(* Logix 5000 project; controller PLC_MCC1300_75F1 vendor 1 type 14 code 166 rev 32.11; software revision 32.04; part 79 of 83 *)
(* tags used below, declared in another part *)
   AUX_xInitialize : BOOL;
   GP_NetDiag : GP_NetworkDiag;
   GP_OB_InitializeDiag : GP_OB_Initialize;
   GP_OB_InitializeDiag_STC : GP_OB_Initialize_STC;
   GP_OB_InitializeMain : GP_OB_Initialize;
   M302SpeedUp : MAC_SpeedUp;
   M307A_M1_DR : AXIS_CIP_DRIVE;
   M307A_M2_DR : AXIS_CIP_DRIVE;
   M307A_M3_DR : AXIS_CIP_DRIVE;
   M351_ALM : MAC_Conveyor_ALM;
   M352_ALM : MAC_Conveyor_ALM;
   M353_ALM : MAC_Conveyor_ALM;
   MCC1300_rgtDiagModule_HMI : GP_NetworkDiag_v1[90];
   TMP_dDirection : DINT;
   TMP_dTarget : DINT;
   TMP_rAcc : REAL;
   TMP_rDec : REAL;
   TMP_rSpeed : REAL;
   Z300_Conveyor : UDT_StandConv[29];
   Z300_Conveyor_IN_MOTION : MAC_Conveyor_ZC_IN_MOTION[29];
   Z300_Conveyor_OUT_MOTION : MAC_Conveyor_ZC_OUT_MOTION[29];
   Z301 : MAC_Zone_ML;
   Z900 : MAC_Zone;
   Z900_HMR : MAC_Zone_HMR;
   Z900_HMW : MAC_Zone_HMW;
(* MainProgram, continued *)

   // #####_HMI_STATUSES_#####
   40: NOP();
   41: XIC(Z900.ST_xZoneError)OTE(Z900_HMR.xZoneAlarm);
   42: XIC(Z900.ST_xCleaningAccepted)OTE(Z900_HMR.xCleaningEnabled);
   43: [MOV(0,Z900_HMR.dCabinetState1) ,[XIC(M351_ALM.rgxStoppingFault_M[0].1) ,XIC(M352_ALM.rgxStoppingFault_M[0].1) ,XIC(M353_ALM.rgxStoppingFault_M[0].1) ] MOV(2,Z900_HMR.dCabinetState1) ,XIC(Z301.OUTPUT_xMCCSafetyLamp) MOV(1,Z900_HMR.dCabinetState1) ];
   44: [XIC(Z900.ST_xManualModeAccepted) MOV(1,Z900_HMR.dZoneMode) ,XIC(Z900.ST_xAutoModeAccepted) MOV(4,Z900_HMR.dZoneMode) ,XIC(Z900.ST_xManualModeRequest) MOV(8,Z900_HMR.dZoneMode) ];
   45: [MOV(2,Z900_HMR.dZoneState) ,XIC(Z900.ST_xStartCycleRequest) XIO(Z900.ST_xCycleON) MOV(4,Z900_HMR.dZoneState) ,XIC(Z900.ST_xCycleON) MOV(1,Z900_HMR.dZoneState) ,XIC(Z900.ST_xStopCycleRequest) MOV(8,Z900_HMR.dZoneState) ,XIO(Z301.INPUT_xMainEmergencyON) MOV(1024,Z900_HMR.dZoneState) ];
   46: [XIC(Z900.ST_xCleaningAccepted) MOV(1,Z900_HMR.dCleaningState) ,XIO(Z900.ST_xCleaningAccepted) MOV(2,Z900_HMR.dCleaningState) ,XIC(Z900.ST_xReqCleaning) XIO(Z900.ST_xCleaningAccepted) MOV(4,Z900_HMR.dCleaningState) ];
   47: [XIC(Z900_HMW.rgxMan.0) OTE(Z900_HMR.rgxMan.0) ,XIC(Z900_HMW.rgxMan.1) OTE(Z900_HMR.rgxMan.1) ];
END_ROUTINE
END_PROGRAM

PROGRAM Modules   (* main routine Main *)

ROUTINE Main   (* ladder *)
   0: GP_OB_Initialize(GP_OB_InitializeDiag,GP_OB_InitializeDiag_STC,AUX_xInitialize);
   1: GP_NetworkDiag(GP_NetDiag,GP_OB_InitializeDiag,ETH_MCC1300,MCC1300_rgtDiagModule_HMI[0]);
   2: GP_NetworkDiag(GP_NetDiag,GP_OB_InitializeDiag,ETH_M2,MCC1300_rgtDiagModule_HMI[1]);
   3: GP_NetworkDiag(GP_NetDiag,GP_OB_InitializeDiag,TD5680AP1,MCC1300_rgtDiagModule_HMI[5]);
   4: GP_NetworkDiag(GP_NetDiag,GP_OB_InitializeDiag,M3683AP1,MCC1300_rgtDiagModule_HMI[6]);
   5: GP_NetworkDiag(GP_NetDiag,GP_OB_InitializeDiag,E152AP1,MCC1300_rgtDiagModule_HMI[7]);
   6: GP_NetworkDiag(GP_NetDiag,GP_OB_InitializeDiag,RIOM13,MCC1300_rgtDiagModule_HMI[8]);
   7: GP_NetworkDiag(GP_NetDiag,GP_OB_InitializeDiag,M3AZ01,MCC1300_rgtDiagModule_HMI[11]);
   8: GP_NetworkDiag(GP_NetDiag,GP_OB_InitializeDiag,M3AZ02,MCC1300_rgtDiagModule_HMI[12]);
   9: GP_NetworkDiag(GP_NetDiag,GP_OB_InitializeDiag,M3AZ03,MCC1300_rgtDiagModule_HMI[13]);
   10: GP_NetworkDiag(GP_NetDiag,GP_OB_InitializeDiag,M3AZ04,MCC1300_rgtDiagModule_HMI[14]);
   11: GP_NetworkDiag(GP_NetDiag,GP_OB_InitializeDiag,M3AZ05,MCC1300_rgtDiagModule_HMI[15]);
   12: GP_NetworkDiag(GP_NetDiag,GP_OB_InitializeDiag,M3AZ06,MCC1300_rgtDiagModule_HMI[16]);
   13: GP_NetworkDiag(GP_NetDiag,GP_OB_InitializeDiag,M3AZ07,MCC1300_rgtDiagModule_HMI[17]);
   14: GP_NetworkDiag(GP_NetDiag,GP_OB_InitializeDiag,M3AZ08,MCC1300_rgtDiagModule_HMI[18]);
   15: GP_NetworkDiag(GP_NetDiag,GP_OB_InitializeDiag,M3AZ09,MCC1300_rgtDiagModule_HMI[19]);
   16: GP_NetworkDiag(GP_NetDiag,GP_OB_InitializeDiag,M3AZ10,MCC1300_rgtDiagModule_HMI[20]);
   17: GP_NetworkDiag(GP_NetDiag,GP_OB_InitializeDiag,TDKAZ00N,MCC1300_rgtDiagModule_HMI[21]);
   18: GP_NetworkDiag(GP_NetDiag,GP_OB_InitializeDiag,TDKAZ00S,MCC1300_rgtDiagModule_HMI[22]);
   19: GP_NetworkDiag(GP_NetDiag,GP_OB_InitializeDiag,TDKAZ01N,MCC1300_rgtDiagModule_HMI[23]);
   20: GP_NetworkDiag(GP_NetDiag,GP_OB_InitializeDiag,TDKAZ01S,MCC1300_rgtDiagModule_HMI[24]);
   21: GP_NetworkDiag(GP_NetDiag,GP_OB_InitializeDiag,TDKAZ02N,MCC1300_rgtDiagModule_HMI[25]);
   22: GP_NetworkDiag(GP_NetDiag,GP_OB_InitializeDiag,TDKAZ02S,MCC1300_rgtDiagModule_HMI[26]);
   23: GP_NetworkDiag(GP_NetDiag,GP_OB_InitializeDiag,TDKAZ03N,MCC1300_rgtDiagModule_HMI[27]);
   24: GP_NetworkDiag(GP_NetDiag,GP_OB_InitializeDiag,TDKAZ03S,MCC1300_rgtDiagModule_HMI[28]);
   25: GP_NetworkDiag(GP_NetDiag,GP_OB_InitializeDiag,TDKAZ04N,MCC1300_rgtDiagModule_HMI[29]);
   26: GP_NetworkDiag(GP_NetDiag,GP_OB_InitializeDiag,TDKAZ04S,MCC1300_rgtDiagModule_HMI[30]);
   27: GP_NetworkDiag(GP_NetDiag,GP_OB_InitializeDiag,TDKAZ05N,MCC1300_rgtDiagModule_HMI[31]);
   28: GP_NetworkDiag(GP_NetDiag,GP_OB_InitializeDiag,TDKAZ05S,MCC1300_rgtDiagModule_HMI[32]);
   29: GP_NetworkDiag(GP_NetDiag,GP_OB_InitializeDiag,TDAZ00N,MCC1300_rgtDiagModule_HMI[33]);
   30: GP_NetworkDiag(GP_NetDiag,GP_OB_InitializeDiag,TDAZ00S,MCC1300_rgtDiagModule_HMI[34]);
   31: GP_NetworkDiag(GP_NetDiag,GP_OB_InitializeDiag,TDAZ01N,MCC1300_rgtDiagModule_HMI[35]);
   32: GP_NetworkDiag(GP_NetDiag,GP_OB_InitializeDiag,TDAZ01S,MCC1300_rgtDiagModule_HMI[36]);
   33: GP_NetworkDiag(GP_NetDiag,GP_OB_InitializeDiag,TDAZ02N,MCC1300_rgtDiagModule_HMI[37]);
   34: GP_NetworkDiag(GP_NetDiag,GP_OB_InitializeDiag,TDAZ02S,MCC1300_rgtDiagModule_HMI[38]);
   35: GP_NetworkDiag(GP_NetDiag,GP_OB_InitializeDiag,TDAZ03N,MCC1300_rgtDiagModule_HMI[39]);
   36: GP_NetworkDiag(GP_NetDiag,GP_OB_InitializeDiag,TDAZ03S,MCC1300_rgtDiagModule_HMI[40]);
   37: GP_NetworkDiag(GP_NetDiag,GP_OB_InitializeDiag,TDAZ04N,MCC1300_rgtDiagModule_HMI[41]);
   38: GP_NetworkDiag(GP_NetDiag,GP_OB_InitializeDiag,TDAZ04S,MCC1300_rgtDiagModule_HMI[42]);
   39: GP_NetworkDiag(GP_NetDiag,GP_OB_InitializeDiag,TDAZ05N,MCC1300_rgtDiagModule_HMI[43]);
   40: GP_NetworkDiag(GP_NetDiag,GP_OB_InitializeDiag,TDAZ05S,MCC1300_rgtDiagModule_HMI[44]);
   41: GP_NetworkDiag(GP_NetDiag,GP_OB_InitializeDiag,D010M1PM1,MCC1300_rgtDiagModule_HMI[46]);
   42: GP_NetworkDiag(GP_NetDiag,GP_OB_InitializeDiag,D010M2PM1,MCC1300_rgtDiagModule_HMI[47]);
   43: GP_NetworkDiag(GP_NetDiag,GP_OB_InitializeDiag,D020M1PM1,MCC1300_rgtDiagModule_HMI[48]);
   44: GP_NetworkDiag(GP_NetDiag,GP_OB_InitializeDiag,E53AZ1,MCC1300_rgtDiagModule_HMI[50]);
   45: GP_NetworkDiag(GP_NetDiag,GP_OB_InitializeDiag,E61AZ1,MCC1300_rgtDiagModule_HMI[51]);
   46: GP_NetworkDiag(GP_NetDiag,GP_OB_InitializeDiag,E62AZ1,MCC1300_rgtDiagModule_HMI[52]);
   47: GP_NetworkDiag(GP_NetDiag,GP_OB_InitializeDiag,E63AZ1,MCC1300_rgtDiagModule_HMI[53]);
   48: GP_NetworkDiag(GP_NetDiag,GP_OB_InitializeDiag,E64AZ1,MCC1300_rgtDiagModule_HMI[54]);
   49: GP_NetworkDiag(GP_NetDiag,GP_OB_InitializeDiag,E65AZ1,MCC1300_rgtDiagModule_HMI[55]);
   50: GP_NetworkDiag(GP_NetDiag,GP_OB_InitializeDiag,E66AZ1,MCC1300_rgtDiagModule_HMI[56]);
   51: GP_NetworkDiag(GP_NetDiag,GP_OB_InitializeDiag,E67AZ1,MCC1300_rgtDiagModule_HMI[57]);
   52: GP_NetworkDiag(GP_NetDiag,GP_OB_InitializeDiag,E71AZ1,MCC1300_rgtDiagModule_HMI[58]);
   53: GP_NetworkDiag(GP_NetDiag,GP_OB_InitializeDiag,E73AZ1,MCC1300_rgtDiagModule_HMI[59]);
   54: GP_NetworkDiag(GP_NetDiag,GP_OB_InitializeDiag,E76AZ1,MCC1300_rgtDiagModule_HMI[60]);
   55: GP_NetworkDiag(GP_NetDiag,GP_OB_InitializeDiag,E77AZ1,MCC1300_rgtDiagModule_HMI[61]);
   56: GP_NetworkDiag(GP_NetDiag,GP_OB_InitializeDiag,E78AZ1,MCC1300_rgtDiagModule_HMI[62]);
   57: GP_NetworkDiag(GP_NetDiag,GP_OB_InitializeDiag,E81AZ1,MCC1300_rgtDiagModule_HMI[63]);
   58: GP_NetworkDiag(GP_NetDiag,GP_OB_InitializeDiag,E82AZ1,MCC1300_rgtDiagModule_HMI[64]);
   59: GP_NetworkDiag(GP_NetDiag,GP_OB_InitializeDiag,E83AZ1,MCC1300_rgtDiagModule_HMI[65]);
   60: GP_NetworkDiag(GP_NetDiag,GP_OB_InitializeDiag,E84AZ1,MCC1300_rgtDiagModule_HMI[66]);
   61: GP_NetworkDiag(GP_NetDiag,GP_OB_InitializeDiag,E85AZ1,MCC1300_rgtDiagModule_HMI[67]);
   62: GP_NetworkDiag(GP_NetDiag,GP_OB_InitializeDiag,E86AZ1,MCC1300_rgtDiagModule_HMI[68]);
   63: GP_NetworkDiag(GP_NetDiag,GP_OB_InitializeDiag,E87AZ1,MCC1300_rgtDiagModule_HMI[69]);
   64: GP_NetworkDiag(GP_NetDiag,GP_OB_InitializeDiag,E88AZ1,MCC1300_rgtDiagModule_HMI[70]);
   65: GP_NetworkDiag(GP_NetDiag,GP_OB_InitializeDiag,E91AZ1,MCC1300_rgtDiagModule_HMI[71]);
   66: GP_NetworkDiag(GP_NetDiag,GP_OB_InitializeDiag,E93AZ1,MCC1300_rgtDiagModule_HMI[72]);
   67: GP_NetworkDiag(GP_NetDiag,GP_OB_InitializeDiag,E96AZ1,MCC1300_rgtDiagModule_HMI[73]);
   68: GP_NetworkDiag(GP_NetDiag,GP_OB_InitializeDiag,E97AZ1,MCC1300_rgtDiagModule_HMI[74]);
   69: GP_NetworkDiag(GP_NetDiag,GP_OB_InitializeDiag,E98AZ1,MCC1300_rgtDiagModule_HMI[75]);
END_ROUTINE
END_PROGRAM

PROGRAM MotionLogic   (* main routine Main *)

ROUTINE M307A_Motion   (* ladder *)
   // M307AM1
   0: NOP();
   1: XIC(Z300_Conveyor[12].OUTPUT_xDriveReset.0)MASR(M307A_M1_DR,Z300_Conveyor_OUT_MOTION[12].DR_MASR_M[0]);
   2: [XIC(Z300_Conveyor[12].OUTPUT_xDriveEnable.[0]) XIO(Z300_Conveyor_OUT_MOTION[12].DR_MSO_M[0].ER) MSO(M307A_M1_DR,Z300_Conveyor_OUT_MOTION[12].DR_MSO_M[0]) ,XIO(Z300_Conveyor_OUT_MOTION[12].DR_MSO_M[0].EN) OTU(Z300_Conveyor_OUT_MOTION[12].DR_MSO_M[0].ER) ,XIO(Z300_Conveyor[12].OUTPUT_xDriveEnable.[0]) OTU(Z300_Conveyor_OUT_MOTION[12].DR_MSO_M[0].EN) XIO(Z300_Conveyor_OUT_MOTION[12].DR_MSF_M[0].ER) MSF(M307A_M1_DR,Z300_Conveyor_OUT_MOTION[12].DR_MSF_M[0]) ,XIO(Z300_Conveyor_OUT_MOTION[12].DR_MSF_M[0].EN) OTU(Z300_Conveyor_OUT_MOTION[12].DR_MSF_M[0].ER) ];
   3: MUL(Z300_Conveyor[12].AUX_rgrAcc_m_s2[0],1000,TMP_rAcc)MUL(Z300_Conveyor[12].AUX_rgrDec_m_s2[0],1000,TMP_rDec)DIV(Z300_Conveyor[12].AUX_rgdRequestSpeed_mm_min[0],60,TMP_rSpeed);
   4: XIC(Z300_Conveyor[12].OS_xStartCount.0)OTU(Z300_Conveyor_IN_MOTION[12].DR_MAR_M[0].PC)OTU(Z300_Conveyor_IN_MOTION[12].DR_MRP_M[0].DN);
   5: [XIC(Z300_Conveyor[12].OUTPUT_xRun.0) MOV(0,TMP_dDirection) ,XIC(Z300_Conveyor[12].OUTPUT_xReverse.0) MOV(1,TMP_dDirection) ][XIO(Z300_Conveyor_IN_MOTION[12].DR_MAR_M[0].PC) ,XIO(Z300_Conveyor_IN_MOTION[12].DR_MRP_M[0].DN) ,XIO(Z300_Conveyor[12].OUTPUT_xPositioning.0) ]MAJ(M307A_M1_DR,Z300_Conveyor_OUT_MOTION[12].DR_MAJ_M[0],TMP_dDirection,TMP_rSpeed,Units per sec,TMP_rAcc,Units per sec2,TMP_rDec,Units per sec2,Trapezoidal,TMP_rAcc,TMP_rDec,Units per sec3,Enabled,Programmed,0,None);
   6: XIC(Z300_Conveyor[12].OS_xStartCount.0)MRP(M307A_M1_DR,Z300_Conveyor_OUT_MOTION[12].DR_MRP_M[0],Absolute,Actual,0);
   7: [XIC(Z300_Conveyor_IN_MOTION[12].DR_MRP_M[0].DN) XIC(Z300_Conveyor[12].OUTPUT_xPositioning.0) [XIC(Z300_Conveyor[12].tmON_PhFilter[0].DN) ,XIC(Z300_Conveyor_IN_MOTION[12].DR_MAR_M[0].EN) ] MAR(M307A_M1_DR,Z300_Conveyor_OUT_MOTION[12].DR_MAR_M[0],Negative_Edge,Disabled,0,0,1) ,XIO(Z300_Conveyor[12].OUTPUT_xPositioning.0) MDR(M307A_M1_DR,Z300_Conveyor_OUT_MOTION[12].DR_MDR_M[0],1) ];
   8: XIC(Z300_Conveyor[12].OUTPUT_xPositioning.0)XIC(Z300_Conveyor_IN_MOTION[12].DR_MAR_M[0].PC)DIV(Z300_Conveyor[12].AUX_rgdTarget_cmm[0],100,TMP_dTarget)ADD(TMP_dTarget,M307A_M1_DR.Registration1Position,TMP_dTarget)MAM(M307A_M1_DR,Z300_Conveyor_OUT_MOTION[12].DR_MAM_M[0],0,TMP_dTarget,TMP_rSpeed,Units per sec,TMP_rAcc,Units per sec2,TMP_rDec,Units per sec2,Trapezoidal,TMP_rAcc,TMP_rDec,Units per sec3,Enabled,Programmed,0,None,0,0);
   9: [XIC(Z300_Conveyor[12].OUTPUT_xChangeSpeed.0) ,XIC(M302SpeedUp.OS_xChangeAccDec) ,XIC(GP_OB_InitializeMain.OUT_xOs_200ms) ][XIO(Z300_Conveyor[12].OUTPUT_xReverse.0) ,XIC(Z300_Conveyor[12].OUTPUT_xReverse.0) MUL(TMP_rSpeed,-1.0,TMP_rSpeed) ]MCD(M307A_M1_DR,Z300_Conveyor_OUT_MOTION[12].DR_MCD_M[0],Jog,Yes,TMP_rSpeed,Yes,TMP_rAcc,Yes,TMP_rDec,No,TMP_rAcc,No,TMP_rDec,Units per sec,Units per sec2,Units per sec2,Units per sec3);
   10: XIO(Z300_Conveyor[12].OUTPUT_xRun.0)XIO(Z300_Conveyor[12].OUTPUT_xReverse.0)[XIC(Z300_Conveyor_IN_MOTION[12].DR_MAJ_M[0].IP) MAS(M307A_M1_DR,Z300_Conveyor_OUT_MOTION[12].DR_MASjog_M[0],Jog,Yes,TMP_rDec,Units per sec2,No,TMP_rDec,Units per sec3) ,XIC(Z300_Conveyor_IN_MOTION[12].DR_MAM_M[0].IP) MAS(M307A_M1_DR,Z300_Conveyor_OUT_MOTION[12].DR_MASpos_M[0],Move,Yes,TMP_rDec,Units per sec2,No,TMP_rDec,Units per sec3) ,XIO(Z300_Conveyor_IN_MOTION[12].DR_MAJ_M[0].IP) XIO(Z300_Conveyor_IN_MOTION[12].DR_MAM_M[0].IP) XIO(Z300_Conveyor_IN_MOTION[12].DR_MASjog_M[0].IP) XIO(Z300_Conveyor_IN_MOTION[12].DR_MASpos_M[0].IP) MAS(M307A_M1_DR,Z300_Conveyor_OUT_MOTION[12].DR_MASall_M[0],All,Yes,TMP_rDec,Units per sec2,No,TMP_rDec,Units per sec3) ];
   // M307AM2
   11: NOP();
   12: XIC(Z300_Conveyor[13].OUTPUT_xDriveReset.0)MASR(M307A_M2_DR,Z300_Conveyor_OUT_MOTION[13].DR_MASR_M[0]);
   13: [XIC(Z300_Conveyor[13].OUTPUT_xDriveEnable.[0]) XIO(Z300_Conveyor_OUT_MOTION[13].DR_MSO_M[0].ER) MSO(M307A_M2_DR,Z300_Conveyor_OUT_MOTION[13].DR_MSO_M[0]) ,XIO(Z300_Conveyor_OUT_MOTION[13].DR_MSO_M[0].EN) OTU(Z300_Conveyor_OUT_MOTION[13].DR_MSO_M[0].ER) ,XIO(Z300_Conveyor[13].OUTPUT_xDriveEnable.[0]) OTU(Z300_Conveyor_OUT_MOTION[13].DR_MSO_M[0].EN) XIO(Z300_Conveyor_OUT_MOTION[13].DR_MSF_M[0].ER) MSF(M307A_M2_DR,Z300_Conveyor_OUT_MOTION[13].DR_MSF_M[0]) ,XIO(Z300_Conveyor_OUT_MOTION[13].DR_MSF_M[0].EN) OTU(Z300_Conveyor_OUT_MOTION[13].DR_MSF_M[0].ER) ];
   14: MUL(Z300_Conveyor[13].AUX_rgrAcc_m_s2[0],1000,TMP_rAcc)MUL(Z300_Conveyor[13].AUX_rgrDec_m_s2[0],1000,TMP_rDec)DIV(Z300_Conveyor[13].AUX_rgdRequestSpeed_mm_min[0],60,TMP_rSpeed);
   15: XIC(Z300_Conveyor[13].OS_xStartCount.0)OTU(Z300_Conveyor_IN_MOTION[13].DR_MAR_M[0].PC)OTU(Z300_Conveyor_IN_MOTION[13].DR_MRP_M[0].DN);
   16: [XIC(Z300_Conveyor[13].OUTPUT_xRun.0) MOV(0,TMP_dDirection) ,XIC(Z300_Conveyor[13].OUTPUT_xReverse.0) MOV(1,TMP_dDirection) ][XIO(Z300_Conveyor_IN_MOTION[13].DR_MAR_M[0].PC) ,XIO(Z300_Conveyor_IN_MOTION[13].DR_MRP_M[0].DN) ,XIO(Z300_Conveyor[13].OUTPUT_xPositioning.0) ]MAJ(M307A_M2_DR,Z300_Conveyor_OUT_MOTION[13].DR_MAJ_M[0],TMP_dDirection,TMP_rSpeed,Units per sec,TMP_rAcc,Units per sec2,TMP_rDec,Units per sec2,Trapezoidal,TMP_rAcc,TMP_rDec,Units per sec3,Enabled,Programmed,0,None);
   17: XIC(Z300_Conveyor[13].OS_xStartCount.0)MRP(M307A_M2_DR,Z300_Conveyor_OUT_MOTION[13].DR_MRP_M[0],Absolute,Actual,0);
   18: [XIC(Z300_Conveyor_IN_MOTION[13].DR_MRP_M[0].DN) XIC(Z300_Conveyor[13].OUTPUT_xPositioning.0) [XIC(Z300_Conveyor[13].tmON_PhFilter[0].DN) ,XIC(Z300_Conveyor_IN_MOTION[13].DR_MAR_M[0].EN) ] MAR(M307A_M2_DR,Z300_Conveyor_OUT_MOTION[13].DR_MAR_M[0],Negative_Edge,Disabled,0,0,1) ,XIO(Z300_Conveyor[13].OUTPUT_xPositioning.0) MDR(M307A_M2_DR,Z300_Conveyor_OUT_MOTION[13].DR_MDR_M[0],1) ];
   19: XIC(Z300_Conveyor[13].OUTPUT_xPositioning.0)XIC(Z300_Conveyor_IN_MOTION[13].DR_MAR_M[0].PC)DIV(Z300_Conveyor[13].AUX_rgdTarget_cmm[0],100,TMP_dTarget)ADD(TMP_dTarget,M307A_M2_DR.Registration1Position,TMP_dTarget)MAM(M307A_M2_DR,Z300_Conveyor_OUT_MOTION[13].DR_MAM_M[0],0,TMP_dTarget,TMP_rSpeed,Units per sec,TMP_rAcc,Units per sec2,TMP_rDec,Units per sec2,Trapezoidal,TMP_rAcc,TMP_rDec,Units per sec3,Enabled,Programmed,0,None,0,0);
   20: [XIC(Z300_Conveyor[13].OUTPUT_xChangeSpeed.0) ,XIC(M302SpeedUp.OS_xChangeAccDec) ,XIC(GP_OB_InitializeMain.OUT_xOs_200ms) ][XIO(Z300_Conveyor[13].OUTPUT_xReverse.0) ,XIC(Z300_Conveyor[13].OUTPUT_xReverse.0) MUL(TMP_rSpeed,-1.0,TMP_rSpeed) ]MCD(M307A_M2_DR,Z300_Conveyor_OUT_MOTION[13].DR_MCD_M[0],Jog,Yes,TMP_rSpeed,Yes,TMP_rAcc,Yes,TMP_rDec,No,TMP_rAcc,No,TMP_rDec,Units per sec,Units per sec2,Units per sec2,Units per sec3);
   21: XIO(Z300_Conveyor[13].OUTPUT_xRun.0)XIO(Z300_Conveyor[13].OUTPUT_xReverse.0)[XIC(Z300_Conveyor_IN_MOTION[13].DR_MAJ_M[0].IP) MAS(M307A_M2_DR,Z300_Conveyor_OUT_MOTION[13].DR_MASjog_M[0],Jog,Yes,TMP_rDec,Units per sec2,No,TMP_rDec,Units per sec3) ,XIC(Z300_Conveyor_IN_MOTION[13].DR_MAM_M[0].IP) MAS(M307A_M2_DR,Z300_Conveyor_OUT_MOTION[13].DR_MASpos_M[0],Move,Yes,TMP_rDec,Units per sec2,No,TMP_rDec,Units per sec3) ,XIO(Z300_Conveyor_IN_MOTION[13].DR_MAJ_M[0].IP) XIO(Z300_Conveyor_IN_MOTION[13].DR_MAM_M[0].IP) XIO(Z300_Conveyor_IN_MOTION[13].DR_MASjog_M[0].IP) XIO(Z300_Conveyor_IN_MOTION[13].DR_MASpos_M[0].IP) MAS(M307A_M2_DR,Z300_Conveyor_OUT_MOTION[13].DR_MASall_M[0],All,Yes,TMP_rDec,Units per sec2,No,TMP_rDec,Units per sec3) ];
   // M307AM3
   22: NOP();
   23: XIC(Z300_Conveyor[14].OUTPUT_xDriveReset.0)MASR(M307A_M3_DR,Z300_Conveyor_OUT_MOTION[14].DR_MASR_M[0]);
